REGION Network 14: MFC- 4011:Mass Flow Controller Flow for Calcination
   RUNG wire#powerrail
      "MFC-4011-F_DB"(EnableHighAlarms := wire#w1, EnableLowAlarms := wire#w2, Mode := 2, RAIVI :=, RAIVR :=, "TI Fail" :=, SAI =>)
   END_RUNG
   RUNG wire#powerrail
      Contact( "R-401_DB".Equipments.Valves."FV-4011".Enable )
      { S7_Templates := "SrcType := Int" } GT_Contact(in1 := "R-401_DB".Status."Step", in2 := 23)
   END_RUNG wire#w1
   RUNG wire#powerrail
      Contact( "R-401_DB".Equipments.Valves."FV-4011".Enable )
      { S7_Templates := "SrcType := Int" } GT_Contact(in1 := "R-401_DB".Status."Step", in2 := 23)
   END_RUNG wire#w2
   RUNG wire#powerrail
      I_Contact( false )
      { S7_GenerateENO := "TRUE" } Move(in := "MFC-4011_MB_R_DB".MB_Data.Buffer[4], out1 => "MFC-4011-F_DB".RAIVR)
   END_RUNG
   // the same network as SCL:
   "MFC-4011-F_DB"(Mode := 2,   // "TX-AI"
                   EnableHighAlarms := "R-401_DB".Equipments.Valves."FV-4011".Enable AND ("R-401_DB".Status."Step" > 23),
                   EnableLowAlarms := "R-401_DB".Equipments.Valves."FV-4011".Enable AND ("R-401_DB".Status."Step" > 23));
   IF NOT false THEN "MFC-4011-F_DB".RAIVR := "MFC-4011_MB_R_DB".MB_Data.Buffer[4]; END_IF;
END_REGION

REGION Network 15: MFC- 4012:Mass Flow Controller Flow for Calcination
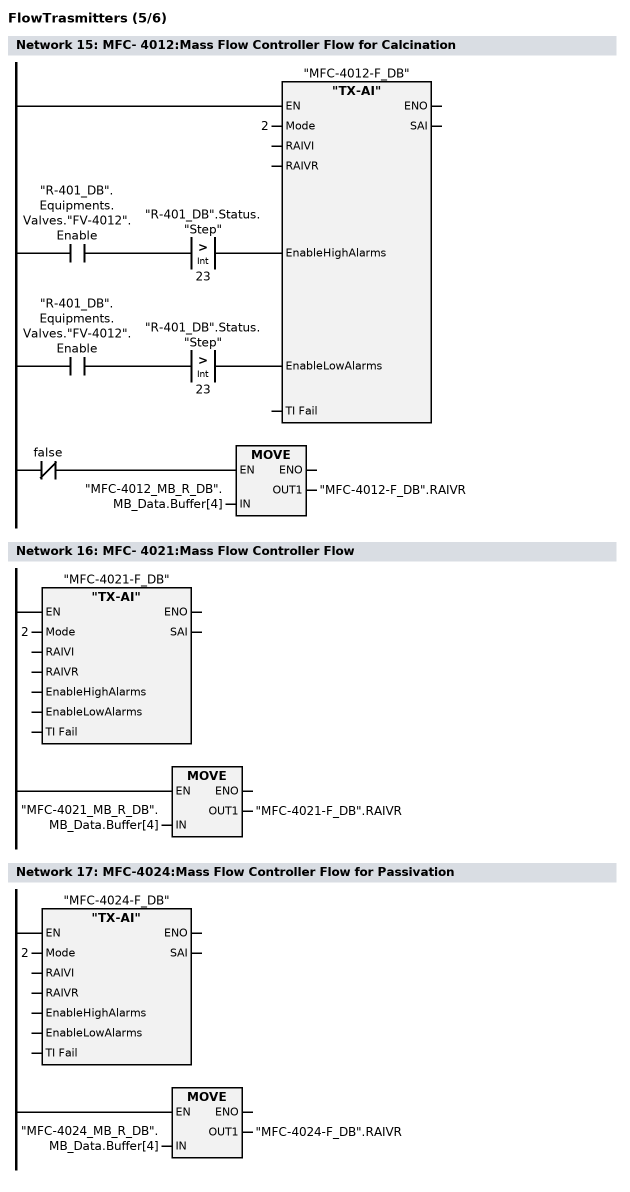
   RUNG wire#powerrail
      "MFC-4012-F_DB"(EnableHighAlarms := wire#w1, EnableLowAlarms := wire#w2, Mode := 2, RAIVI :=, RAIVR :=, "TI Fail" :=, SAI =>)
   END_RUNG
   RUNG wire#powerrail
      Contact( "R-401_DB".Equipments.Valves."FV-4012".Enable )
      { S7_Templates := "SrcType := Int" } GT_Contact(in1 := "R-401_DB".Status."Step", in2 := 23)
   END_RUNG wire#w1
   RUNG wire#powerrail
      Contact( "R-401_DB".Equipments.Valves."FV-4012".Enable )
      { S7_Templates := "SrcType := Int" } GT_Contact(in1 := "R-401_DB".Status."Step", in2 := 23)
   END_RUNG wire#w2
   RUNG wire#powerrail
      I_Contact( false )
      { S7_GenerateENO := "TRUE" } Move(in := "MFC-4012_MB_R_DB".MB_Data.Buffer[4], out1 => "MFC-4012-F_DB".RAIVR)
   END_RUNG
   // the same network as SCL:
   "MFC-4012-F_DB"(Mode := 2,   // "TX-AI"
                   EnableHighAlarms := "R-401_DB".Equipments.Valves."FV-4012".Enable AND ("R-401_DB".Status."Step" > 23),
                   EnableLowAlarms := "R-401_DB".Equipments.Valves."FV-4012".Enable AND ("R-401_DB".Status."Step" > 23));
   IF NOT false THEN "MFC-4012-F_DB".RAIVR := "MFC-4012_MB_R_DB".MB_Data.Buffer[4]; END_IF;
END_REGION

REGION Network 16: MFC- 4021:Mass Flow Controller Flow
   RUNG wire#powerrail
      "MFC-4021-F_DB"(Mode := 2, RAIVI :=, RAIVR :=, EnableHighAlarms :=, EnableLowAlarms :=, "TI Fail" :=, SAI =>)
   END_RUNG
   RUNG wire#powerrail
      { S7_GenerateENO := "TRUE" } Move(in := "MFC-4021_MB_R_DB".MB_Data.Buffer[4], out1 => "MFC-4021-F_DB".RAIVR)
   END_RUNG
   // the same network as SCL:
   "MFC-4021-F_DB"(Mode := 2);   // "TX-AI"
   "MFC-4021-F_DB".RAIVR := "MFC-4021_MB_R_DB".MB_Data.Buffer[4];
END_REGION

REGION Network 17: MFC-4024:Mass Flow Controller Flow for Passivation
   RUNG wire#powerrail
      "MFC-4024-F_DB"(Mode := 2, RAIVI :=, RAIVR :=, EnableHighAlarms :=, EnableLowAlarms :=, "TI Fail" :=, SAI =>)
   END_RUNG
   RUNG wire#powerrail
      { S7_GenerateENO := "TRUE" } Move(in := "MFC-4024_MB_R_DB".MB_Data.Buffer[4], out1 => "MFC-4024-F_DB".RAIVR)
   END_RUNG
   // the same network as SCL:
   "MFC-4024-F_DB"(Mode := 2);   // "TX-AI"
   "MFC-4024-F_DB".RAIVR := "MFC-4024_MB_R_DB".MB_Data.Buffer[4];
END_REGION

REGION Network 18: MFC-4025:Mass Flow Controller Flow for Passivation
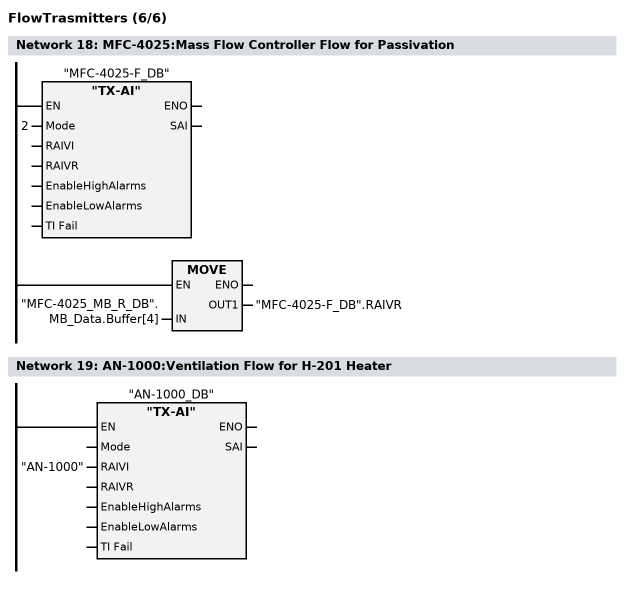
   RUNG wire#powerrail
      "MFC-4025-F_DB"(Mode := 2, RAIVI :=, RAIVR :=, EnableHighAlarms :=, EnableLowAlarms :=, "TI Fail" :=, SAI =>)
   END_RUNG
   RUNG wire#powerrail
      { S7_GenerateENO := "TRUE" } Move(in := "MFC-4025_MB_R_DB".MB_Data.Buffer[4], out1 => "MFC-4025-F_DB".RAIVR)
   END_RUNG
   // the same network as SCL:
   "MFC-4025-F_DB"(Mode := 2);   // "TX-AI"
   "MFC-4025-F_DB".RAIVR := "MFC-4025_MB_R_DB".MB_Data.Buffer[4];
END_REGION

REGION Network 19: AN-1000:Ventilation Flow for H-201 Heater
   RUNG wire#powerrail
      "AN-1000_DB"(Mode :=, RAIVI := "AN-1000", RAIVR :=, EnableHighAlarms :=, EnableLowAlarms :=, "TI Fail" :=, SAI =>)
   END_RUNG
   // the same network as SCL:
   "AN-1000_DB"(RAIVI := "AN-1000");   // "TX-AI"
END_REGION
END_FUNCTION

// folder: Analogs inputs/Trasmitters/Hydrogen Gas Trasmitters

FUNCTION "HydrogenGasTrasmitters" : Void   // FC17, LAD
TITLE = Hydrogen Gas Detector Trasmitters
{ S7_Optimized_Access := 'TRUE' }
VERSION : 0.1
// Updated Date:
// Note:
BEGIN

REGION Network 1: GD-H2-1: Hydrogen Gas Detector #1
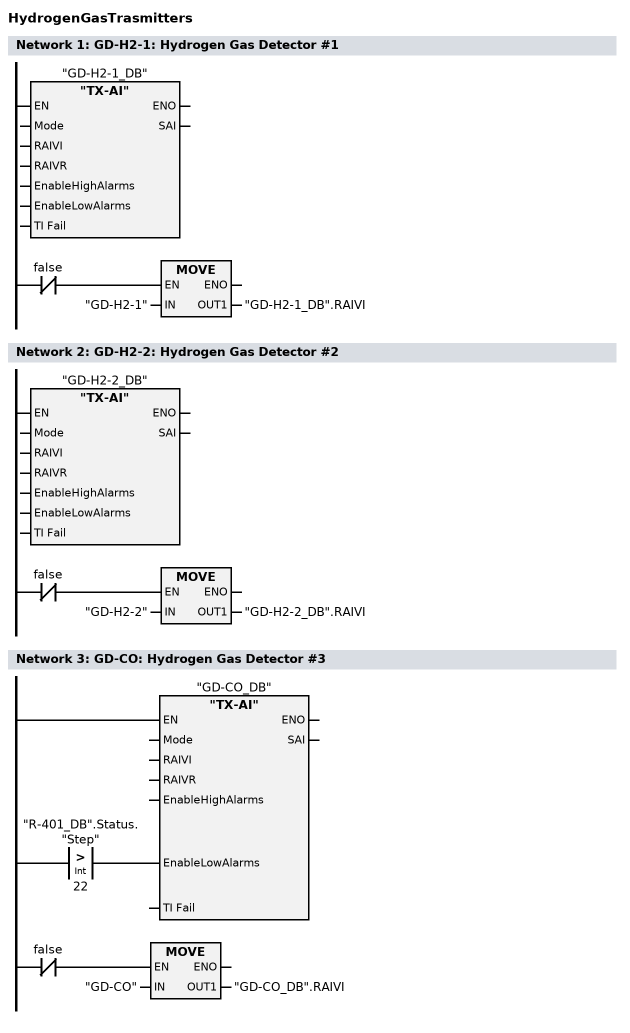
   RUNG wire#powerrail
      "GD-H2-1_DB"(Mode :=, RAIVI :=, RAIVR :=, EnableHighAlarms :=, EnableLowAlarms :=, "TI Fail" :=, SAI =>)
   END_RUNG
   RUNG wire#powerrail
      I_Contact( false )
      { S7_GenerateENO := "TRUE" } Move(in := "GD-H2-1", out1 => "GD-H2-1_DB".RAIVI)
   END_RUNG
   // the same network as SCL:
   "GD-H2-1_DB"();   // "TX-AI"
   IF NOT false THEN "GD-H2-1_DB".RAIVI := "GD-H2-1"; END_IF;
END_REGION

REGION Network 2: GD-H2-2: Hydrogen Gas Detector #2
   RUNG wire#powerrail
      "GD-H2-2_DB"(Mode :=, RAIVI :=, RAIVR :=, EnableHighAlarms :=, EnableLowAlarms :=, "TI Fail" :=, SAI =>)
   END_RUNG
   RUNG wire#powerrail
      I_Contact( false )
      { S7_GenerateENO := "TRUE" } Move(in := "GD-H2-2", out1 => "GD-H2-2_DB".RAIVI)
   END_RUNG
   // the same network as SCL:
   "GD-H2-2_DB"();   // "TX-AI"
   IF NOT false THEN "GD-H2-2_DB".RAIVI := "GD-H2-2"; END_IF;
END_REGION

REGION Network 3: GD-CO: Hydrogen Gas Detector #3
   RUNG wire#powerrail
      "GD-CO_DB"(EnableLowAlarms := wire#w1, Mode :=, RAIVI :=, RAIVR :=, EnableHighAlarms :=, "TI Fail" :=, SAI =>)
   END_RUNG
   RUNG wire#powerrail
      { S7_Templates := "SrcType := Int" } GT_Contact(in1 := "R-401_DB".Status."Step", in2 := 22)
   END_RUNG wire#w1
   RUNG wire#powerrail
      I_Contact( false )
      { S7_GenerateENO := "TRUE" } Move(in := "GD-CO", out1 => "GD-CO_DB".RAIVI)
   END_RUNG
   // the same network as SCL:
   "GD-CO_DB"(EnableLowAlarms := "R-401_DB".Status."Step" > 22);   // "TX-AI"
   IF NOT false THEN "GD-CO_DB".RAIVI := "GD-CO"; END_IF;
END_REGION
END_FUNCTION

// folder: Analogs inputs/Trasmitters/Level Trasmitters

FUNCTION "LevelTrasmitters" : Void   // FC11, LAD
{ S7_Optimized_Access := 'TRUE' }
VERSION : 0.1
// Updated Date:
// Note:
   VAR_TEMP
      "LT-1011_Vol_Gal" : Real;
      "LT-1021_Vol_Gal" : Real;
      "LT-101_h" : Real;
      "LT-102_h" : Real;
   END_VAR
BEGIN

REGION Network 1: LT-1011 : T-101 X Material Level
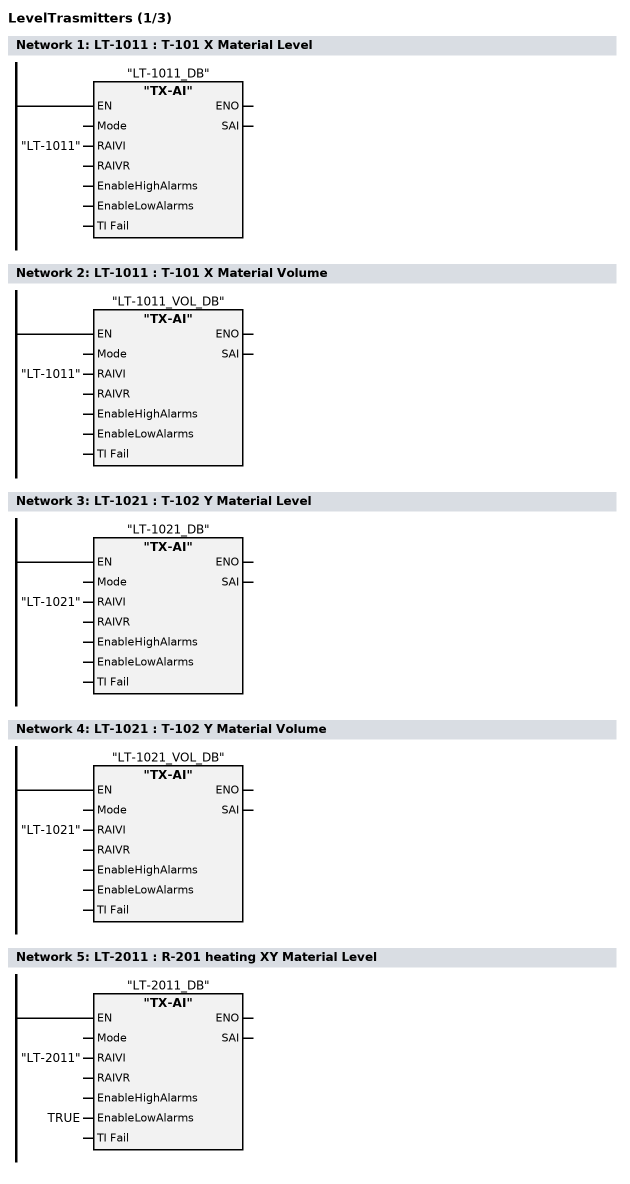
   RUNG wire#powerrail
      "LT-1011_DB"(Mode :=, RAIVI := "LT-1011", RAIVR :=, EnableHighAlarms :=, EnableLowAlarms :=, "TI Fail" :=, SAI =>)
   END_RUNG
   // the same network as SCL:
   "LT-1011_DB"(RAIVI := "LT-1011");   // "TX-AI"
END_REGION

REGION Network 2: LT-1011 : T-101 X Material Volume
   RUNG wire#powerrail
      "LT-1011_VOL_DB"(Mode :=, RAIVI := "LT-1011", RAIVR :=, EnableHighAlarms :=, EnableLowAlarms :=, "TI Fail" :=, SAI =>)
   END_RUNG
   // the same network as SCL:
   "LT-1011_VOL_DB"(RAIVI := "LT-1011");   // "TX-AI"
END_REGION

REGION Network 3: LT-1021 : T-102 Y Material Level
   RUNG wire#powerrail
      "LT-1021_DB"(Mode :=, RAIVI := "LT-1021", RAIVR :=, EnableHighAlarms :=, EnableLowAlarms :=, "TI Fail" :=, SAI =>)
   END_RUNG
   // the same network as SCL:
   "LT-1021_DB"(RAIVI := "LT-1021");   // "TX-AI"
END_REGION

REGION Network 4: LT-1021 : T-102 Y Material Volume
   RUNG wire#powerrail
      "LT-1021_VOL_DB"(Mode :=, RAIVI := "LT-1021", RAIVR :=, EnableHighAlarms :=, EnableLowAlarms :=, "TI Fail" :=, SAI =>)
   END_RUNG
   // the same network as SCL:
   "LT-1021_VOL_DB"(RAIVI := "LT-1021");   // "TX-AI"
END_REGION

REGION Network 5: LT-2011 : R-201 heating XY Material Level
   RUNG wire#powerrail
      "LT-2011_DB"(Mode :=, RAIVI := "LT-2011", RAIVR :=, EnableHighAlarms :=, EnableLowAlarms := TRUE, "TI Fail" :=, SAI =>)
   END_RUNG
   // the same network as SCL:
   "LT-2011_DB"(RAIVI := "LT-2011", EnableLowAlarms := TRUE);   // "TX-AI"
END_REGION

REGION Network 6: LT-2011 : R-201 heating XY Material Volume
   // Max Volume: 200.0 Liters
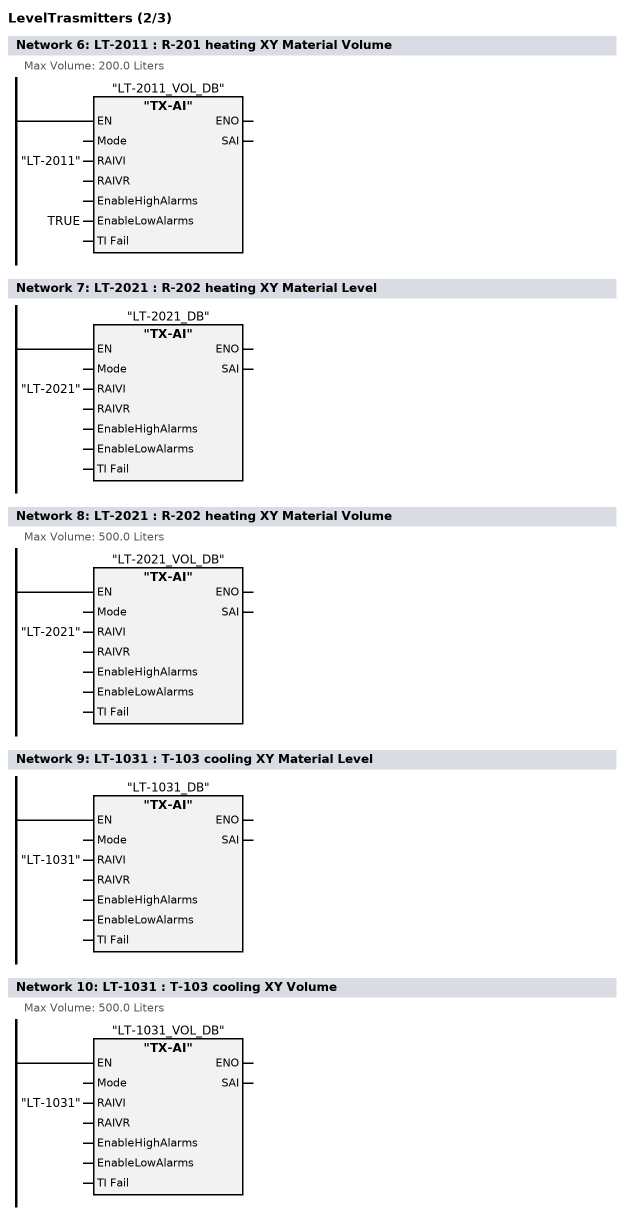
   RUNG wire#powerrail
      "LT-2011_VOL_DB"(Mode :=, RAIVI := "LT-2011", RAIVR :=, EnableHighAlarms :=, EnableLowAlarms := TRUE, "TI Fail" :=, SAI =>)
   END_RUNG
   // the same network as SCL:
   "LT-2011_VOL_DB"(RAIVI := "LT-2011", EnableLowAlarms := TRUE);   // "TX-AI"
END_REGION

REGION Network 7: LT-2021 : R-202 heating XY Material Level
   RUNG wire#powerrail
      "LT-2021_DB"(Mode :=, RAIVI := "LT-2021", RAIVR :=, EnableHighAlarms :=, EnableLowAlarms :=, "TI Fail" :=, SAI =>)
   END_RUNG
   // the same network as SCL:
   "LT-2021_DB"(RAIVI := "LT-2021");   // "TX-AI"
END_REGION

REGION Network 8: LT-2021 : R-202 heating XY Material Volume
   // Max Volume: 500.0 Liters
   RUNG wire#powerrail
      "LT-2021_VOL_DB"(Mode :=, RAIVI := "LT-2021", RAIVR :=, EnableHighAlarms :=, EnableLowAlarms :=, "TI Fail" :=, SAI =>)
   END_RUNG
   // the same network as SCL:
   "LT-2021_VOL_DB"(RAIVI := "LT-2021");   // "TX-AI"
END_REGION

REGION Network 9: LT-1031 : T-103 cooling XY Material Level
   RUNG wire#powerrail
      "LT-1031_DB"(Mode :=, RAIVI := "LT-1031", RAIVR :=, EnableHighAlarms :=, EnableLowAlarms :=, "TI Fail" :=, SAI =>)
   END_RUNG
   // the same network as SCL:
   "LT-1031_DB"(RAIVI := "LT-1031");   // "TX-AI"
END_REGION

REGION Network 10: LT-1031 : T-103 cooling XY Volume
   // Max Volume: 500.0 Liters
   RUNG wire#powerrail
      "LT-1031_VOL_DB"(Mode :=, RAIVI := "LT-1031", RAIVR :=, EnableHighAlarms :=, EnableLowAlarms :=, "TI Fail" :=, SAI =>)
   END_RUNG
   // the same network as SCL:
   "LT-1031_VOL_DB"(RAIVI := "LT-1031");   // "TX-AI"
END_REGION

REGION Network 11: LT-1051 : T-105 Centrifuge wastewater Level
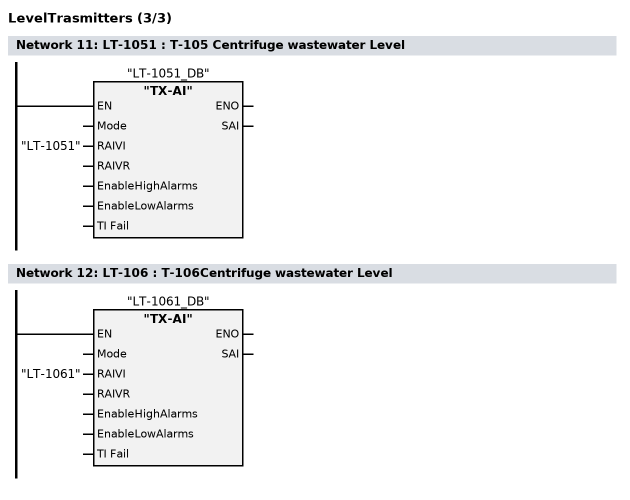
   RUNG wire#powerrail
      "LT-1051_DB"(Mode :=, RAIVI := "LT-1051", RAIVR :=, EnableHighAlarms :=, EnableLowAlarms :=, "TI Fail" :=, SAI =>)
   END_RUNG
   // the same network as SCL:
   "LT-1051_DB"(RAIVI := "LT-1051");   // "TX-AI"
END_REGION

REGION Network 12: LT-106 : T-106Centrifuge wastewater Level
   RUNG wire#powerrail
      "LT-1061_DB"(Mode :=, RAIVI := "LT-1061", RAIVR :=, EnableHighAlarms :=, EnableLowAlarms :=, "TI Fail" :=, SAI =>)
   END_RUNG
   // the same network as SCL:
   "LT-1061_DB"(RAIVI := "LT-1061");   // "TX-AI"
END_REGION
END_FUNCTION

// folder: Analogs inputs/Trasmitters/Ph Trasmitters

FUNCTION "PhTrasmitters" : Void   // FC15, LAD
{ S7_Optimized_Access := 'TRUE' }
VERSION : 0.1
BEGIN

REGION Network 1: pH-2011 : R-201 pH #1
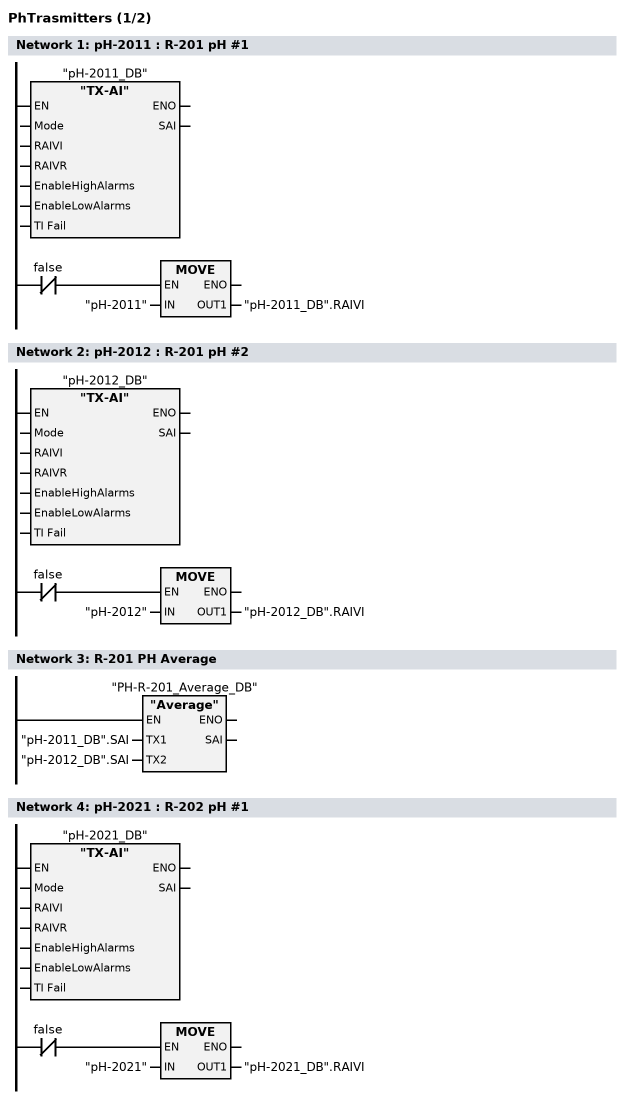
   RUNG wire#powerrail
      "pH-2011_DB"(Mode :=, RAIVI :=, RAIVR :=, EnableHighAlarms :=, EnableLowAlarms :=, "TI Fail" :=, SAI =>)
   END_RUNG
   RUNG wire#powerrail
      I_Contact( false )
      { S7_GenerateENO := "TRUE" } Move(in := "pH-2011", out1 => "pH-2011_DB".RAIVI)
   END_RUNG
   // the same network as SCL:
   "pH-2011_DB"();   // "TX-AI"
   IF NOT false THEN "pH-2011_DB".RAIVI := "pH-2011"; END_IF;
END_REGION

REGION Network 2: pH-2012 : R-201 pH #2
   RUNG wire#powerrail
      "pH-2012_DB"(Mode :=, RAIVI :=, RAIVR :=, EnableHighAlarms :=, EnableLowAlarms :=, "TI Fail" :=, SAI =>)
   END_RUNG
   RUNG wire#powerrail
      I_Contact( false )
      { S7_GenerateENO := "TRUE" } Move(in := "pH-2012", out1 => "pH-2012_DB".RAIVI)
   END_RUNG
   // the same network as SCL:
   "pH-2012_DB"();   // "TX-AI"
   IF NOT false THEN "pH-2012_DB".RAIVI := "pH-2012"; END_IF;
END_REGION

REGION Network 3: R-201 PH Average
   RUNG wire#powerrail
      "PH-R-201_Average_DB"(TX1 := "pH-2011_DB".SAI, TX2 := "pH-2012_DB".SAI, SAI =>)
   END_RUNG
   // the same network as SCL:
   "PH-R-201_Average_DB"(TX1 := "pH-2011_DB".SAI, TX2 := "pH-2012_DB".SAI);   // "Average"
END_REGION

REGION Network 4: pH-2021 : R-202 pH #1
   RUNG wire#powerrail
      "pH-2021_DB"(Mode :=, RAIVI :=, RAIVR :=, EnableHighAlarms :=, EnableLowAlarms :=, "TI Fail" :=, SAI =>)
   END_RUNG
   RUNG wire#powerrail
      I_Contact( false )
      { S7_GenerateENO := "TRUE" } Move(in := "pH-2021", out1 => "pH-2021_DB".RAIVI)
   END_RUNG
   // the same network as SCL:
   "pH-2021_DB"();   // "TX-AI"
   IF NOT false THEN "pH-2021_DB".RAIVI := "pH-2021"; END_IF;
END_REGION

REGION Network 5: pH-2022 : R-202 pH #2
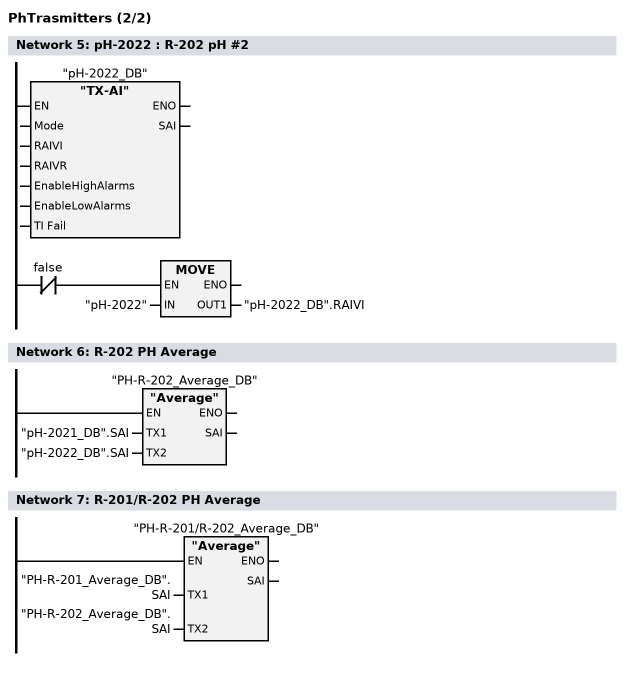
   RUNG wire#powerrail
      "pH-2022_DB"(Mode :=, RAIVI :=, RAIVR :=, EnableHighAlarms :=, EnableLowAlarms :=, "TI Fail" :=, SAI =>)
   END_RUNG
   RUNG wire#powerrail
      I_Contact( false )
      { S7_GenerateENO := "TRUE" } Move(in := "pH-2022", out1 => "pH-2022_DB".RAIVI)
   END_RUNG
   // the same network as SCL:
   "pH-2022_DB"();   // "TX-AI"
   IF NOT false THEN "pH-2022_DB".RAIVI := "pH-2022"; END_IF;
END_REGION

REGION Network 6: R-202 PH Average
   RUNG wire#powerrail
      "PH-R-202_Average_DB"(TX1 := "pH-2021_DB".SAI, TX2 := "pH-2022_DB".SAI, SAI =>)
   END_RUNG
   // the same network as SCL:
   "PH-R-202_Average_DB"(TX1 := "pH-2021_DB".SAI, TX2 := "pH-2022_DB".SAI);   // "Average"
END_REGION

REGION Network 7: R-201/R-202 PH Average
   RUNG wire#powerrail
      "PH-R-201/R-202_Average_DB"(TX1 := "PH-R-201_Average_DB".SAI, TX2 := "PH-R-202_Average_DB".SAI, SAI =>)
   END_RUNG
   // the same network as SCL:
   "PH-R-201/R-202_Average_DB"(TX1 := "PH-R-201_Average_DB".SAI, TX2 := "PH-R-202_Average_DB".SAI);   // "Average"
END_REGION
END_FUNCTION

// folder: Analogs inputs/Trasmitters/Pressure Trasmitters

FUNCTION "PressureTrasmitters" : Void   // FC12, LAD
{ S7_Optimized_Access := 'TRUE' }
VERSION : 0.1
BEGIN

REGION Network 1: PRESSURE TX P101A
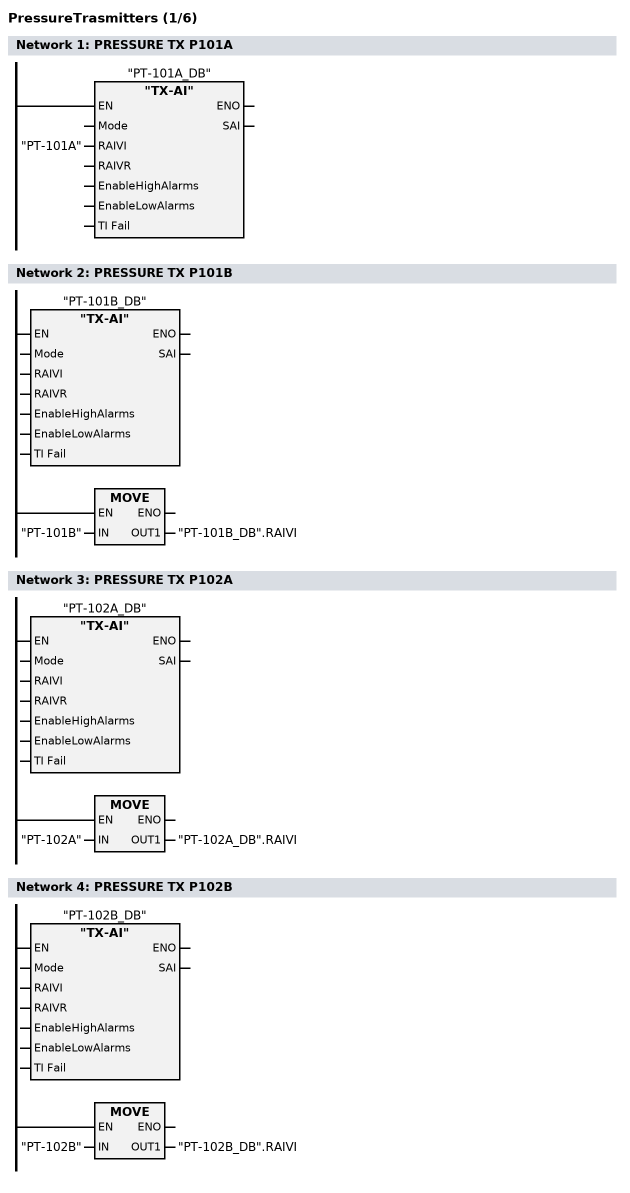
   RUNG wire#powerrail
      "PT-101A_DB"(Mode :=, RAIVI := "PT-101A", RAIVR :=, EnableHighAlarms :=, EnableLowAlarms :=, "TI Fail" :=, SAI =>)
   END_RUNG
   // the same network as SCL:
   "PT-101A_DB"(RAIVI := "PT-101A");   // "TX-AI"
END_REGION

REGION Network 2: PRESSURE TX P101B
   RUNG wire#powerrail
      "PT-101B_DB"(Mode :=, RAIVI :=, RAIVR :=, EnableHighAlarms :=, EnableLowAlarms :=, "TI Fail" :=, SAI =>)
   END_RUNG
   RUNG wire#powerrail
      { S7_GenerateENO := "TRUE" } Move(in := "PT-101B", out1 => "PT-101B_DB".RAIVI)
   END_RUNG
   // the same network as SCL:
   "PT-101B_DB"();   // "TX-AI"
   "PT-101B_DB".RAIVI := "PT-101B";
END_REGION

REGION Network 3: PRESSURE TX P102A
   RUNG wire#powerrail
      "PT-102A_DB"(Mode :=, RAIVI :=, RAIVR :=, EnableHighAlarms :=, EnableLowAlarms :=, "TI Fail" :=, SAI =>)
   END_RUNG
   RUNG wire#powerrail
      { S7_GenerateENO := "TRUE" } Move(in := "PT-102A", out1 => "PT-102A_DB".RAIVI)
   END_RUNG
   // the same network as SCL:
   "PT-102A_DB"();   // "TX-AI"
   "PT-102A_DB".RAIVI := "PT-102A";
END_REGION

REGION Network 4: PRESSURE TX P102B
   RUNG wire#powerrail
      "PT-102B_DB"(Mode :=, RAIVI :=, RAIVR :=, EnableHighAlarms :=, EnableLowAlarms :=, "TI Fail" :=, SAI =>)
   END_RUNG
   RUNG wire#powerrail
      { S7_GenerateENO := "TRUE" } Move(in := "PT-102B", out1 => "PT-102B_DB".RAIVI)
   END_RUNG
   // the same network as SCL:
   "PT-102B_DB"();   // "TX-AI"
   "PT-102B_DB".RAIVI := "PT-102B";
END_REGION

REGION Network 5: PRESSURE TX P103A
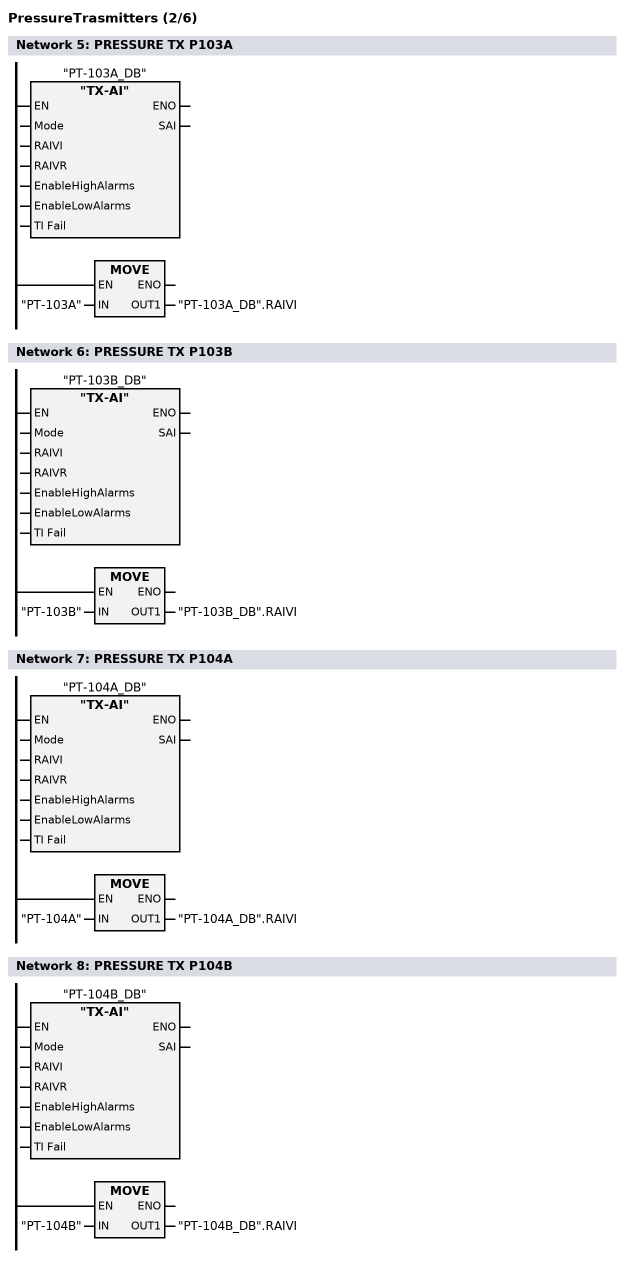
   RUNG wire#powerrail
      "PT-103A_DB"(Mode :=, RAIVI :=, RAIVR :=, EnableHighAlarms :=, EnableLowAlarms :=, "TI Fail" :=, SAI =>)
   END_RUNG
   RUNG wire#powerrail
      { S7_GenerateENO := "TRUE" } Move(in := "PT-103A", out1 => "PT-103A_DB".RAIVI)
   END_RUNG
   // the same network as SCL:
   "PT-103A_DB"();   // "TX-AI"
   "PT-103A_DB".RAIVI := "PT-103A";
END_REGION

REGION Network 6: PRESSURE TX P103B
   RUNG wire#powerrail
      "PT-103B_DB"(Mode :=, RAIVI :=, RAIVR :=, EnableHighAlarms :=, EnableLowAlarms :=, "TI Fail" :=, SAI =>)
   END_RUNG
   RUNG wire#powerrail
      { S7_GenerateENO := "TRUE" } Move(in := "PT-103B", out1 => "PT-103B_DB".RAIVI)
   END_RUNG
   // the same network as SCL:
   "PT-103B_DB"();   // "TX-AI"
   "PT-103B_DB".RAIVI := "PT-103B";
END_REGION

REGION Network 7: PRESSURE TX P104A
   RUNG wire#powerrail
      "PT-104A_DB"(Mode :=, RAIVI :=, RAIVR :=, EnableHighAlarms :=, EnableLowAlarms :=, "TI Fail" :=, SAI =>)
   END_RUNG
   RUNG wire#powerrail
      { S7_GenerateENO := "TRUE" } Move(in := "PT-104A", out1 => "PT-104A_DB".RAIVI)
   END_RUNG
   // the same network as SCL:
   "PT-104A_DB"();   // "TX-AI"
   "PT-104A_DB".RAIVI := "PT-104A";
END_REGION

REGION Network 8: PRESSURE TX P104B
   RUNG wire#powerrail
      "PT-104B_DB"(Mode :=, RAIVI :=, RAIVR :=, EnableHighAlarms :=, EnableLowAlarms :=, "TI Fail" :=, SAI =>)
   END_RUNG
   RUNG wire#powerrail
      { S7_GenerateENO := "TRUE" } Move(in := "PT-104B", out1 => "PT-104B_DB".RAIVI)
   END_RUNG
   // the same network as SCL:
   "PT-104B_DB"();   // "TX-AI"
   "PT-104B_DB".RAIVI := "PT-104B";
END_REGION

REGION Network 9: PRESSURE TX P201A
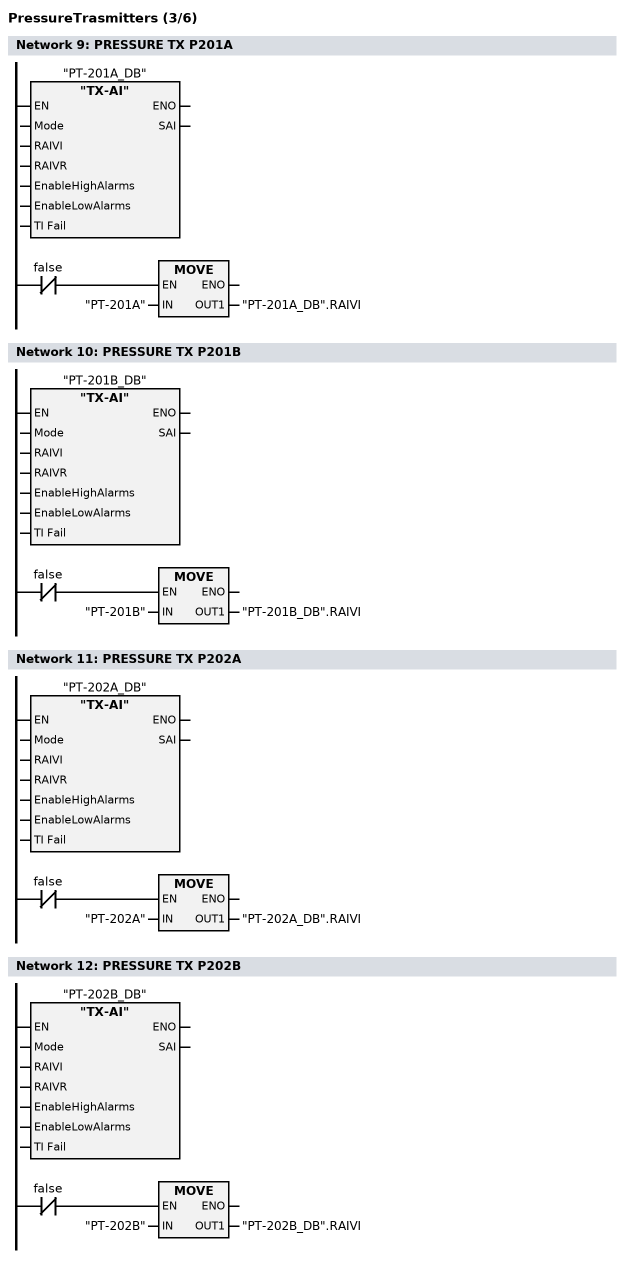
   RUNG wire#powerrail
      "PT-201A_DB"(Mode :=, RAIVI :=, RAIVR :=, EnableHighAlarms :=, EnableLowAlarms :=, "TI Fail" :=, SAI =>)
   END_RUNG
   RUNG wire#powerrail
      I_Contact( false )
      { S7_GenerateENO := "TRUE" } Move(in := "PT-201A", out1 => "PT-201A_DB".RAIVI)
   END_RUNG
   // the same network as SCL:
   "PT-201A_DB"();   // "TX-AI"
   IF NOT false THEN "PT-201A_DB".RAIVI := "PT-201A"; END_IF;
END_REGION

REGION Network 10: PRESSURE TX P201B
   RUNG wire#powerrail
      "PT-201B_DB"(Mode :=, RAIVI :=, RAIVR :=, EnableHighAlarms :=, EnableLowAlarms :=, "TI Fail" :=, SAI =>)
   END_RUNG
   RUNG wire#powerrail
      I_Contact( false )
      { S7_GenerateENO := "TRUE" } Move(in := "PT-201B", out1 => "PT-201B_DB".RAIVI)
   END_RUNG
   // the same network as SCL:
   "PT-201B_DB"();   // "TX-AI"
   IF NOT false THEN "PT-201B_DB".RAIVI := "PT-201B"; END_IF;
END_REGION

REGION Network 11: PRESSURE TX P202A
   RUNG wire#powerrail
      "PT-202A_DB"(Mode :=, RAIVI :=, RAIVR :=, EnableHighAlarms :=, EnableLowAlarms :=, "TI Fail" :=, SAI =>)
   END_RUNG
   RUNG wire#powerrail
      I_Contact( false )
      { S7_GenerateENO := "TRUE" } Move(in := "PT-202A", out1 => "PT-202A_DB".RAIVI)
   END_RUNG
   // the same network as SCL:
   "PT-202A_DB"();   // "TX-AI"
   IF NOT false THEN "PT-202A_DB".RAIVI := "PT-202A"; END_IF;
END_REGION

REGION Network 12: PRESSURE TX P202B
   RUNG wire#powerrail
      "PT-202B_DB"(Mode :=, RAIVI :=, RAIVR :=, EnableHighAlarms :=, EnableLowAlarms :=, "TI Fail" :=, SAI =>)
   END_RUNG
   RUNG wire#powerrail
      I_Contact( false )
      { S7_GenerateENO := "TRUE" } Move(in := "PT-202B", out1 => "PT-202B_DB".RAIVI)
   END_RUNG
   // the same network as SCL:
   "PT-202B_DB"();   // "TX-AI"
   IF NOT false THEN "PT-202B_DB".RAIVI := "PT-202B"; END_IF;
END_REGION

REGION Network 13: PRESSURE TX P301A
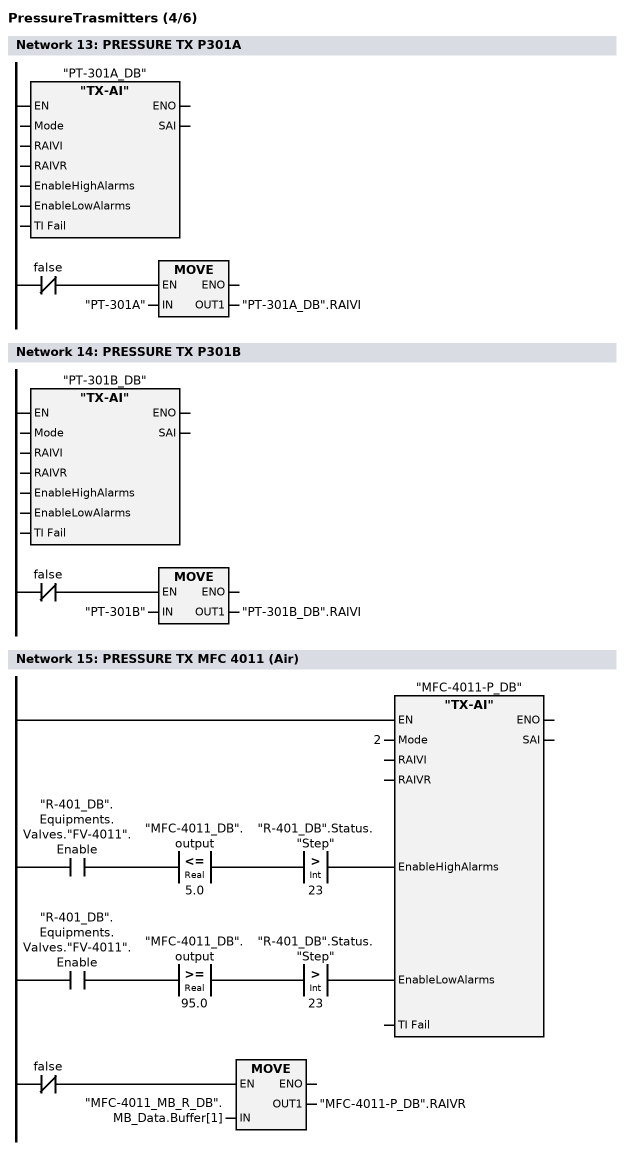
   RUNG wire#powerrail
      "PT-301A_DB"(Mode :=, RAIVI :=, RAIVR :=, EnableHighAlarms :=, EnableLowAlarms :=, "TI Fail" :=, SAI =>)
   END_RUNG
   RUNG wire#powerrail
      I_Contact( false )
      { S7_GenerateENO := "TRUE" } Move(in := "PT-301A", out1 => "PT-301A_DB".RAIVI)
   END_RUNG
   // the same network as SCL:
   "PT-301A_DB"();   // "TX-AI"
   IF NOT false THEN "PT-301A_DB".RAIVI := "PT-301A"; END_IF;
END_REGION

REGION Network 14: PRESSURE TX P301B
   RUNG wire#powerrail
      "PT-301B_DB"(Mode :=, RAIVI :=, RAIVR :=, EnableHighAlarms :=, EnableLowAlarms :=, "TI Fail" :=, SAI =>)
   END_RUNG
   RUNG wire#powerrail
      I_Contact( false )
      { S7_GenerateENO := "TRUE" } Move(in := "PT-301B", out1 => "PT-301B_DB".RAIVI)
   END_RUNG
   // the same network as SCL:
   "PT-301B_DB"();   // "TX-AI"
   IF NOT false THEN "PT-301B_DB".RAIVI := "PT-301B"; END_IF;
END_REGION

REGION Network 15: PRESSURE TX MFC 4011 (Air)
   RUNG wire#powerrail
      "MFC-4011-P_DB"(EnableHighAlarms := wire#w1, EnableLowAlarms := wire#w2, Mode := 2, RAIVI :=, RAIVR :=, "TI Fail" :=, SAI =>)
   END_RUNG
   RUNG wire#powerrail
      Contact( "R-401_DB".Equipments.Valves."FV-4011".Enable )
      { S7_Templates := "SrcType := Real" } LE_Contact(in1 := "MFC-4011_DB".output, in2 := 5.0)
      { S7_Templates := "SrcType := Int" } GT_Contact(in1 := "R-401_DB".Status."Step", in2 := 23)
   END_RUNG wire#w1
   RUNG wire#powerrail
      Contact( "R-401_DB".Equipments.Valves."FV-4011".Enable )
      { S7_Templates := "SrcType := Real" } GE_Contact(in1 := "MFC-4011_DB".output, in2 := 95.0)
      { S7_Templates := "SrcType := Int" } GT_Contact(in1 := "R-401_DB".Status."Step", in2 := 23)
   END_RUNG wire#w2
   RUNG wire#powerrail
      I_Contact( false )
      { S7_GenerateENO := "TRUE" } Move(in := "MFC-4011_MB_R_DB".MB_Data.Buffer[1], out1 => "MFC-4011-P_DB".RAIVR)
   END_RUNG
   // the same network as SCL:
   "MFC-4011-P_DB"(Mode := 2,   // "TX-AI"
                   EnableHighAlarms := "R-401_DB".Equipments.Valves."FV-4011".Enable AND ("MFC-4011_DB".output <= 5.0) AND ("R-401_DB".Status."Step" > 23),
                   EnableLowAlarms := "R-401_DB".Equipments.Valves."FV-4011".Enable AND ("MFC-4011_DB".output >= 95.0) AND ("R-401_DB".Status."Step" > 23));
   IF NOT false THEN "MFC-4011-P_DB".RAIVR := "MFC-4011_MB_R_DB".MB_Data.Buffer[1]; END_IF;
END_REGION

REGION Network 16: PRESSURE TX MFC 4012 ( N2 )
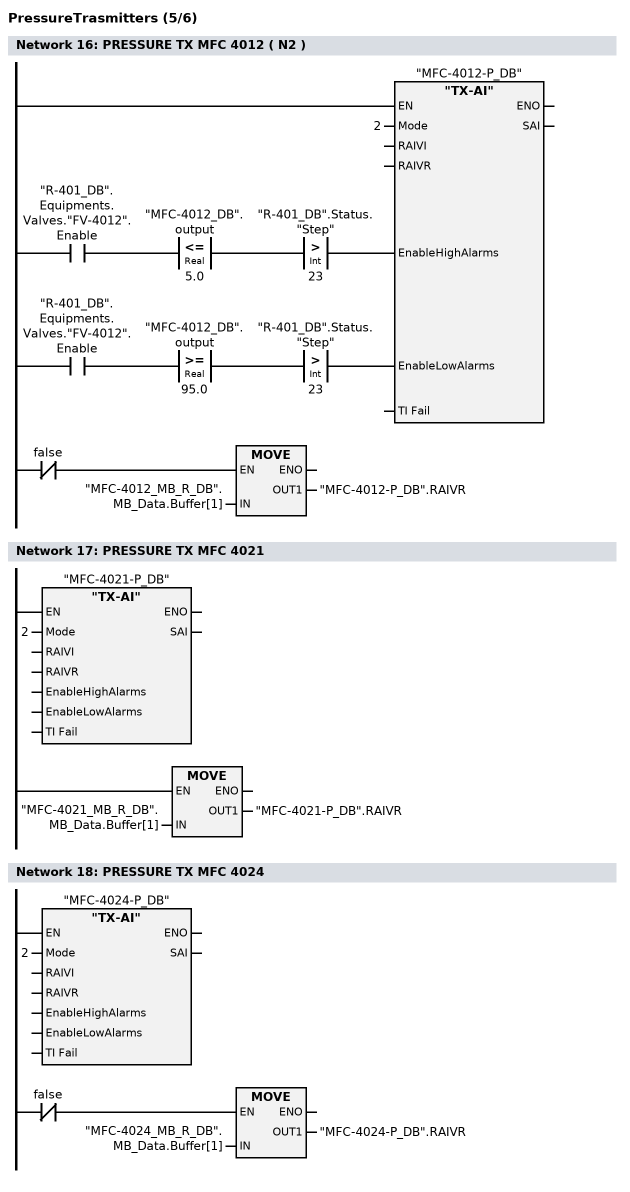
   RUNG wire#powerrail
      "MFC-4012-P_DB"(EnableHighAlarms := wire#w1, EnableLowAlarms := wire#w2, Mode := 2, RAIVI :=, RAIVR :=, "TI Fail" :=, SAI =>)
   END_RUNG
   RUNG wire#powerrail
      Contact( "R-401_DB".Equipments.Valves."FV-4012".Enable )
      { S7_Templates := "SrcType := Real" } LE_Contact(in1 := "MFC-4012_DB".output, in2 := 5.0)
      { S7_Templates := "SrcType := Int" } GT_Contact(in1 := "R-401_DB".Status."Step", in2 := 23)
   END_RUNG wire#w1
   RUNG wire#powerrail
      Contact( "R-401_DB".Equipments.Valves."FV-4012".Enable )
      { S7_Templates := "SrcType := Real" } GE_Contact(in1 := "MFC-4012_DB".output, in2 := 95.0)
      { S7_Templates := "SrcType := Int" } GT_Contact(in1 := "R-401_DB".Status."Step", in2 := 23)
   END_RUNG wire#w2
   RUNG wire#powerrail
      I_Contact( false )
      { S7_GenerateENO := "TRUE" } Move(in := "MFC-4012_MB_R_DB".MB_Data.Buffer[1], out1 => "MFC-4012-P_DB".RAIVR)
   END_RUNG
   // the same network as SCL:
   "MFC-4012-P_DB"(Mode := 2,   // "TX-AI"
                   EnableHighAlarms := "R-401_DB".Equipments.Valves."FV-4012".Enable AND ("MFC-4012_DB".output <= 5.0) AND ("R-401_DB".Status."Step" > 23),
                   EnableLowAlarms := "R-401_DB".Equipments.Valves."FV-4012".Enable AND ("MFC-4012_DB".output >= 95.0) AND ("R-401_DB".Status."Step" > 23));
   IF NOT false THEN "MFC-4012-P_DB".RAIVR := "MFC-4012_MB_R_DB".MB_Data.Buffer[1]; END_IF;
END_REGION

REGION Network 17: PRESSURE TX MFC 4021
   RUNG wire#powerrail
      "MFC-4021-P_DB"(Mode := 2, RAIVI :=, RAIVR :=, EnableHighAlarms :=, EnableLowAlarms :=, "TI Fail" :=, SAI =>)
   END_RUNG
   RUNG wire#powerrail
      { S7_GenerateENO := "TRUE" } Move(in := "MFC-4021_MB_R_DB".MB_Data.Buffer[1], out1 => "MFC-4021-P_DB".RAIVR)
   END_RUNG
   // the same network as SCL:
   "MFC-4021-P_DB"(Mode := 2);   // "TX-AI"
   "MFC-4021-P_DB".RAIVR := "MFC-4021_MB_R_DB".MB_Data.Buffer[1];
END_REGION

REGION Network 18: PRESSURE TX MFC 4024
   RUNG wire#powerrail
      "MFC-4024-P_DB"(Mode := 2, RAIVI :=, RAIVR :=, EnableHighAlarms :=, EnableLowAlarms :=, "TI Fail" :=, SAI =>)
   END_RUNG
   RUNG wire#powerrail
      I_Contact( false )
      { S7_GenerateENO := "TRUE" } Move(in := "MFC-4024_MB_R_DB".MB_Data.Buffer[1], out1 => "MFC-4024-P_DB".RAIVR)
   END_RUNG
   // the same network as SCL:
   "MFC-4024-P_DB"(Mode := 2);   // "TX-AI"
   IF NOT false THEN "MFC-4024-P_DB".RAIVR := "MFC-4024_MB_R_DB".MB_Data.Buffer[1]; END_IF;
END_REGION

REGION Network 19: PRESSURE TX MFC 4025
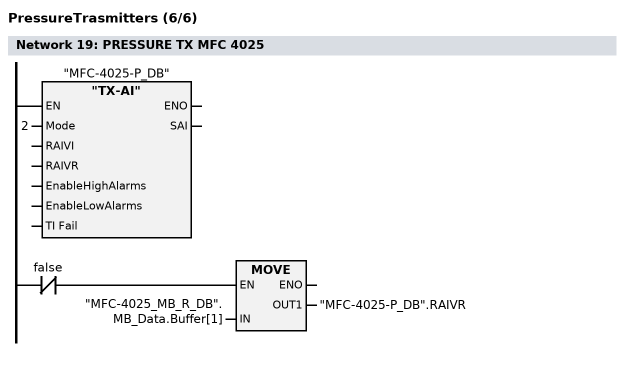
   RUNG wire#powerrail
      "MFC-4025-P_DB"(Mode := 2, RAIVI :=, RAIVR :=, EnableHighAlarms :=, EnableLowAlarms :=, "TI Fail" :=, SAI =>)
   END_RUNG
   RUNG wire#powerrail
      I_Contact( false )
      { S7_GenerateENO := "TRUE" } Move(in := "MFC-4025_MB_R_DB".MB_Data.Buffer[1], out1 => "MFC-4025-P_DB".RAIVR)
   END_RUNG
   // the same network as SCL:
   "MFC-4025-P_DB"(Mode := 2);   // "TX-AI"
   IF NOT false THEN "MFC-4025-P_DB".RAIVR := "MFC-4025_MB_R_DB".MB_Data.Buffer[1]; END_IF;
END_REGION
END_FUNCTION

// folder: Analogs inputs/Trasmitters/Temperature Trasmitters

FUNCTION "TemperatureTrasmitters" : Void   // FC13, LAD
{ S7_Optimized_Access := 'TRUE' }
VERSION : 0.1
BEGIN

REGION Network 1: TT-1031 : T-103 Temperature
